(* Logix 5000 project; controller PLC_MCC1300_75F1 vendor 1 type 14 code 166 rev 32.11; software revision 32.04; part 28 of 83 *)
(* tags used below, declared in another part *)
   AUX_tCapsConveyor_NULL : UDT_CapsConveyor_ZC;
   AUX_xInitialize : BOOL;
   CM_AreaStackerToLine_JS1 : CM_AreaStackerToLine;
   CM_AreaStackerToLine_JS1_Sync : CM_AreaStackerToLine;
   CM_AreaStackerToLine_JS2 : CM_AreaStackerToLine;
   CM_AreaStackerToLine_JS2_Sync : CM_AreaStackerToLine;
   CM_ConveyorStackerToLine_JS1 : CM_ConveyorStackerToLine;
   CM_ConveyorStackerToLine_JS1_Sync : CM_ConveyorStackerToLine;
   CM_ConveyorStackerToLine_JS2 : CM_ConveyorStackerToLine;
   CM_ConveyorStackerToLine_JS2_Sync : CM_ConveyorStackerToLine;
   CM_DATA_Z410_Rx : UDT_PlateData_Convoy;
   CM_DATA_Z410_Rx_Sync : UDT_PlateData_Convoy;
   CM_DATA_Z410_Rx_TmpBuffer : SINT[104];
   CM_DATA_Z410_Tx : UDT_PlateData_Convoy;
   CM_DATA_Z410_Tx_MSG : MESSAGE;
   CM_DATA_Z410_Tx_PH : DINT;
   CM_DATA_Z410_Tx_TempBuffer : SINT[104];
   CM_DATA_Z410_Tx_tmON : TIMER;
   CM_DATA_Z420_Rx : UDT_PlateData_Convoy;
   CM_DATA_Z420_Rx_Sync : UDT_PlateData_Convoy;
   CM_DATA_Z420_Rx_TmpBuffer : SINT[104];
   CM_DATA_Z420_Tx : UDT_PlateData_Convoy;
   CM_DATA_Z420_Tx_MSG : MESSAGE;
   CM_DATA_Z420_Tx_PH : DINT;
   CM_DATA_Z420_Tx_TempBuffer : SINT[104];
   CM_DATA_Z420_Tx_tmON : TIMER;
   CM_LineToAreaStacker_JS1 : CM_LineToAreaStacker;
   CM_LineToAreaStacker_JS2 : CM_LineToAreaStacker;
   CM_LineToConveyorStacker_JS1 : CM_LineToConveyorStacker;
   CM_LineToConveyorStacker_JS2 : CM_LineToConveyorStacker;
   CNV10_FLT : ALIAS FOR I[4].9;
   CNV11_FLT : ALIAS FOR I[4].10;
   CNV12_FLT : ALIAS FOR I[4].11;
   CNV1_FLT : ALIAS FOR I[4].0;
   CNV2_FLT : ALIAS FOR I[4].1;
   CNV3_FLT : ALIAS FOR I[4].2;
   CNV4_FLT : ALIAS FOR I[4].3;
   CNV5_FLT : ALIAS FOR I[4].4;
   CNV6_FLT : ALIAS FOR I[4].5;
   CNV7_FLT : ALIAS FOR I[4].6;
   CNV8_FLT : ALIAS FOR I[4].7;
   CNV9_FLT : ALIAS FOR I[4].8;
   CONST_tPlant : UDT_PLANT_CONSTANTS;
   DROP_NO1_CRSH : ALIAS FOR I[73].12;
   GP_OB_InitializeMain : GP_OB_Initialize;
   GP_OB_InitializeMain_STC : GP_OB_Initialize_STC;
   I : INT[128];   // Local Input Updates Input Slot 2
   M2_DRV_CONT_ON : ALIAS FOR I[2].1;
   M2_DRV_FLT_LMP : ALIAS FOR O[9].0;
   M302SpeedUp : MAC_SpeedUp;
   M307ASpeedUp : MAC_SpeedUp;
   M30xTrimDeck : MAC_TrimmingDeck[5];
   M30xTrimWheel : MAC_TrimmingWheels[5];
   M310Popup : MAC_Popup_ZC[2];
   M310Popup_SL_DATA : UDT_Convoy_SL;
   M312 : MAC_Conveyor_Single;
   M312_SpaceConv_Utilities : SpaceConv_Utilities;
   M315Popup : MAC_Popup_ZC[2];
   M315Popup_SL_DATA : UDT_Convoy_SL;
   M350Popup : MAC_Popup_ZC;
   M410_DATA_xSendERR : BOOL;
   M420_DATA_xSendERR : BOOL;
   N130 : INT[8];
   N131 : INT[8];
   O : INT[128];
   REL_DATARCVD_N : ALIAS FOR O[54].2;
   REL_DATARCVDS : ALIAS FOR O[58].2;
   REL_REJWINLAMPN : ALIAS FOR O[54].3;
   REL_REJWINLAMPS : ALIAS FOR O[58].3;
   T4 : TIMER[51];
   TMP_d : DINT;
   TMP_dIndex : DINT;
   TMP_dIndexCapConv : DINT;
   TMP_dIndexConv : DINT;
   TMP_dLineSize : DINT;
   tony_always_false : BOOL;
   xAlwaysOFF : BOOL;
   Z300_Conveyor : UDT_StandConv[29];
   Z300_Conveyor_Conf : UDT_Conveyor_Config[29];
   Z300_dEndTrackingPosition : DINT;
   Z300_dStartTrackingPosition : DINT;
   Z300_LineTracking : UDT_LINE_TRACKING;
   Z301 : MAC_Zone_ML;
   Z401 : MAC_Zone;
   Z401_HMW : MAC_Zone_HMW;

PROGRAM Communication   (* main routine Main *)

ROUTINE CM_Z410   (* ladder *)
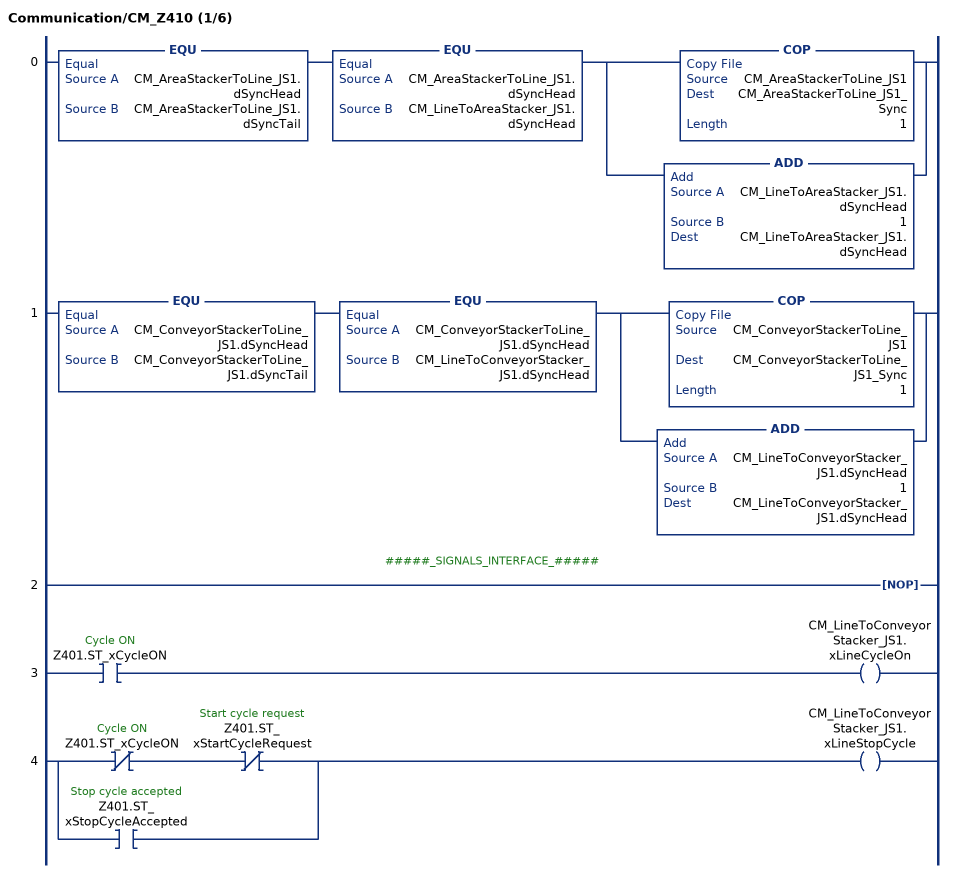
   0: EQU(CM_AreaStackerToLine_JS1.dSyncHead,CM_AreaStackerToLine_JS1.dSyncTail)EQU(CM_AreaStackerToLine_JS1.dSyncHead,CM_LineToAreaStacker_JS1.dSyncHead)[COP(CM_AreaStackerToLine_JS1,CM_AreaStackerToLine_JS1_Sync,1) ,ADD(CM_LineToAreaStacker_JS1.dSyncHead,1,CM_LineToAreaStacker_JS1.dSyncHead) ];
   1: EQU(CM_ConveyorStackerToLine_JS1.dSyncHead,CM_ConveyorStackerToLine_JS1.dSyncTail)EQU(CM_ConveyorStackerToLine_JS1.dSyncHead,CM_LineToConveyorStacker_JS1.dSyncHead)[COP(CM_ConveyorStackerToLine_JS1,CM_ConveyorStackerToLine_JS1_Sync,1) ,ADD(CM_LineToConveyorStacker_JS1.dSyncHead,1,CM_LineToConveyorStacker_JS1.dSyncHead) ];
   // #####_SIGNALS_INTERFACE_#####
   2: NOP();
   3: XIC(Z401.ST_xCycleON)OTE(CM_LineToConveyorStacker_JS1.xLineCycleOn);
   4: [XIO(Z401.ST_xCycleON) XIO(Z401.ST_xStartCycleRequest) ,XIC(Z401.ST_xStopCycleAccepted) ]OTE(CM_LineToConveyorStacker_JS1.xLineStopCycle);
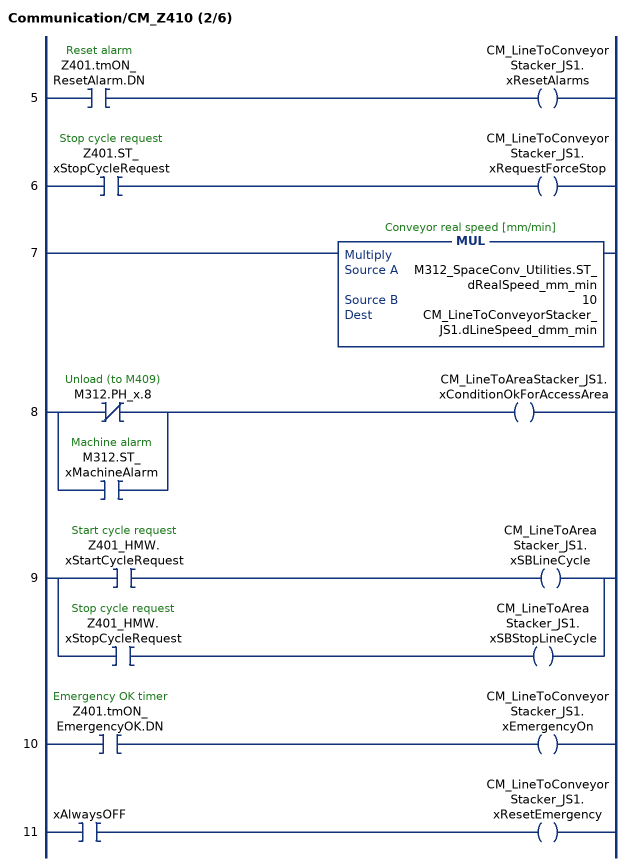
   5: XIC(Z401.tmON_ResetAlarm.DN)OTE(CM_LineToConveyorStacker_JS1.xResetAlarms);
   6: XIC(Z401.ST_xStopCycleRequest)OTE(CM_LineToConveyorStacker_JS1.xRequestForceStop);
   7: MUL(M312_SpaceConv_Utilities.ST_dRealSpeed_mm_min,10,CM_LineToConveyorStacker_JS1.dLineSpeed_dmm_min);
   8: [XIO(M312.PH_x.8) ,XIC(M312.ST_xMachineAlarm) ]OTE(CM_LineToAreaStacker_JS1.xConditionOkForAccessArea);
   9: [XIC(Z401_HMW.xStartCycleRequest) OTE(CM_LineToAreaStacker_JS1.xSBLineCycle) ,XIC(Z401_HMW.xStopCycleRequest) OTE(CM_LineToAreaStacker_JS1.xSBStopLineCycle) ];
   10: XIC(Z401.tmON_EmergencyOK.DN)OTE(CM_LineToConveyorStacker_JS1.xEmergencyOn);
   11: XIC(xAlwaysOFF)OTE(CM_LineToConveyorStacker_JS1.xResetEmergency);
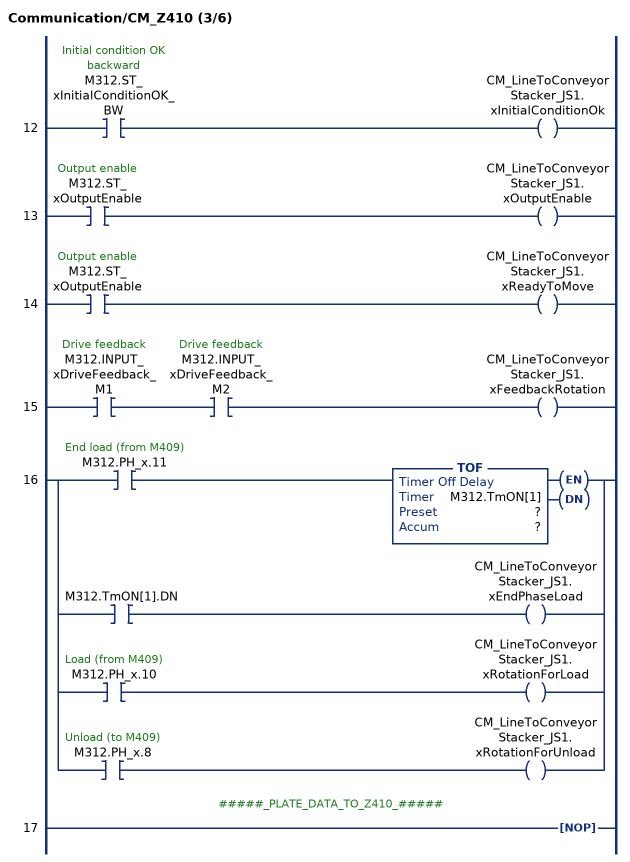
   12: XIC(M312.ST_xInitialConditionOK_BW)OTE(CM_LineToConveyorStacker_JS1.xInitialConditionOk);
   13: XIC(M312.ST_xOutputEnable)OTE(CM_LineToConveyorStacker_JS1.xOutputEnable);
   14: XIC(M312.ST_xOutputEnable)OTE(CM_LineToConveyorStacker_JS1.xReadyToMove);
   15: XIC(M312.INPUT_xDriveFeedback_M1)XIC(M312.INPUT_xDriveFeedback_M2)OTE(CM_LineToConveyorStacker_JS1.xFeedbackRotation);
   16: [[XIC(M312.PH_x.11) TOF(M312.TmON[1],?,?) ,XIC(M312.TmON[1].DN) OTE(CM_LineToConveyorStacker_JS1.xEndPhaseLoad) ] ,XIC(M312.PH_x.10) OTE(CM_LineToConveyorStacker_JS1.xRotationForLoad) ,XIC(M312.PH_x.8) OTE(CM_LineToConveyorStacker_JS1.xRotationForUnload) ];
   // #####_PLATE_DATA_TO_Z410_#####
   17: NOP();
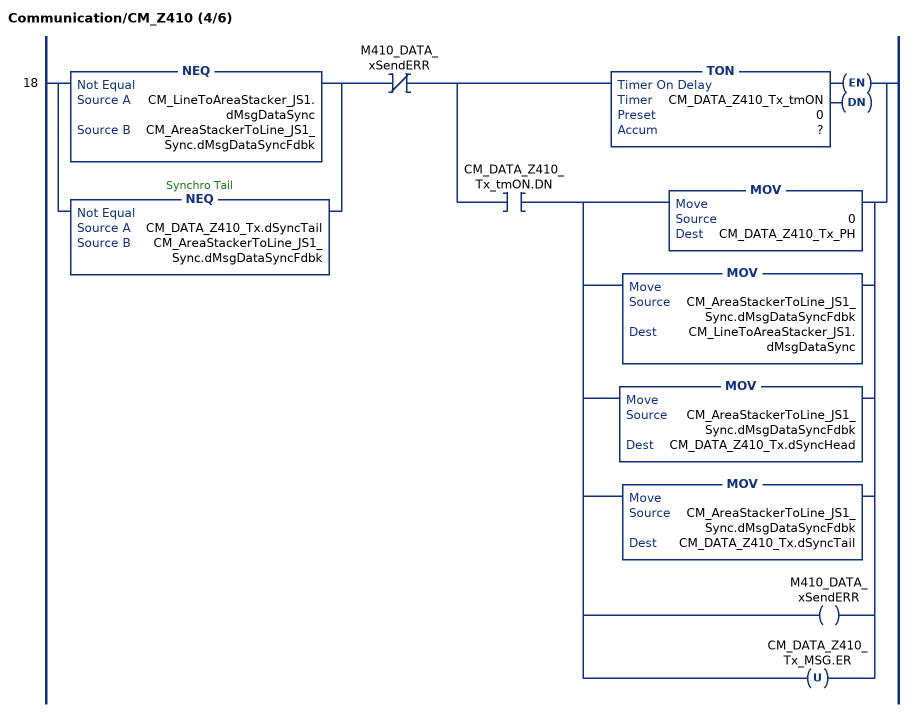
   18: [NEQ(CM_LineToAreaStacker_JS1.dMsgDataSync,CM_AreaStackerToLine_JS1_Sync.dMsgDataSyncFdbk) ,NEQ(CM_DATA_Z410_Tx.dSyncTail,CM_AreaStackerToLine_JS1_Sync.dMsgDataSyncFdbk) ]XIO(M410_DATA_xSendERR)[TON(CM_DATA_Z410_Tx_tmON,?,?) ,XIC(CM_DATA_Z410_Tx_tmON.DN) [MOV(0,CM_DATA_Z410_Tx_PH) ,MOV(CM_AreaStackerToLine_JS1_Sync.dMsgDataSyncFdbk,CM_LineToAreaStacker_JS1.dMsgDataSync) ,MOV(CM_AreaStackerToLine_JS1_Sync.dMsgDataSyncFdbk,CM_DATA_Z410_Tx.dSyncHead) ,MOV(CM_AreaStackerToLine_JS1_Sync.dMsgDataSyncFdbk,CM_DATA_Z410_Tx.dSyncTail) ,OTE(M410_DATA_xSendERR) ,OTU(CM_DATA_Z410_Tx_MSG.ER) ] ];
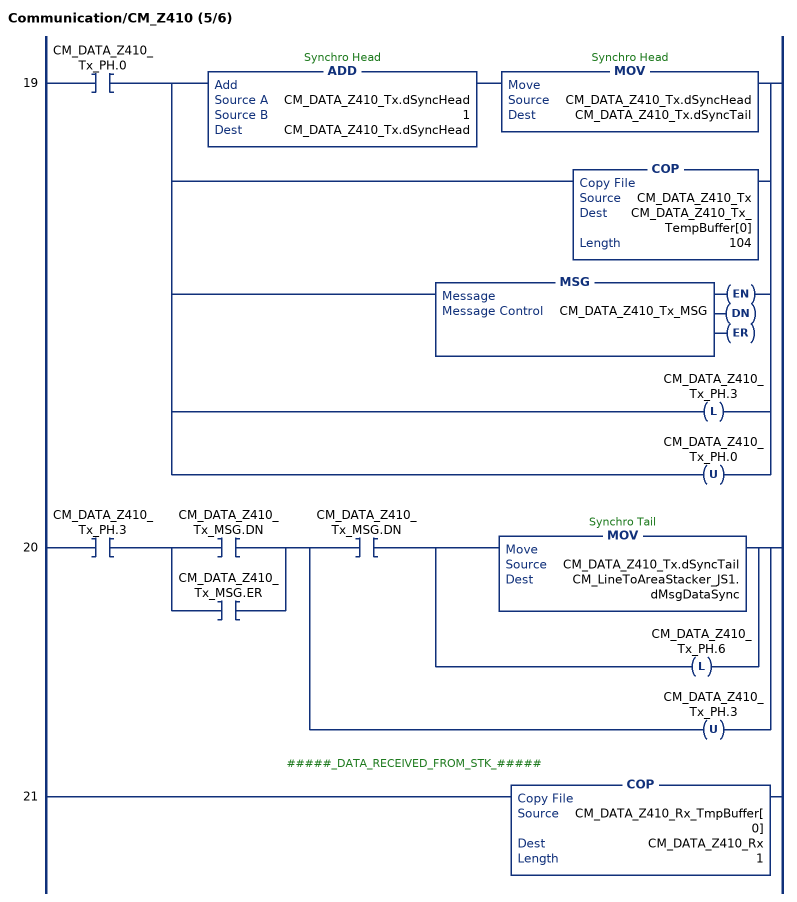
   19: XIC(CM_DATA_Z410_Tx_PH.0)[ADD(CM_DATA_Z410_Tx.dSyncHead,1,CM_DATA_Z410_Tx.dSyncHead) MOV(CM_DATA_Z410_Tx.dSyncHead,CM_DATA_Z410_Tx.dSyncTail) ,COP(CM_DATA_Z410_Tx,CM_DATA_Z410_Tx_TempBuffer[0],104) ,MSG(CM_DATA_Z410_Tx_MSG) ,OTL(CM_DATA_Z410_Tx_PH.3) ,OTU(CM_DATA_Z410_Tx_PH.0) ];
   20: XIC(CM_DATA_Z410_Tx_PH.3)[XIC(CM_DATA_Z410_Tx_MSG.DN) ,XIC(CM_DATA_Z410_Tx_MSG.ER) ][XIC(CM_DATA_Z410_Tx_MSG.DN) [MOV(CM_DATA_Z410_Tx.dSyncTail,CM_LineToAreaStacker_JS1.dMsgDataSync) ,OTL(CM_DATA_Z410_Tx_PH.6) ] ,OTU(CM_DATA_Z410_Tx_PH.3) ];
   // #####_DATA_RECEIVED_FROM_STK_#####
   21: COP(CM_DATA_Z410_Rx_TmpBuffer[0],CM_DATA_Z410_Rx,1);
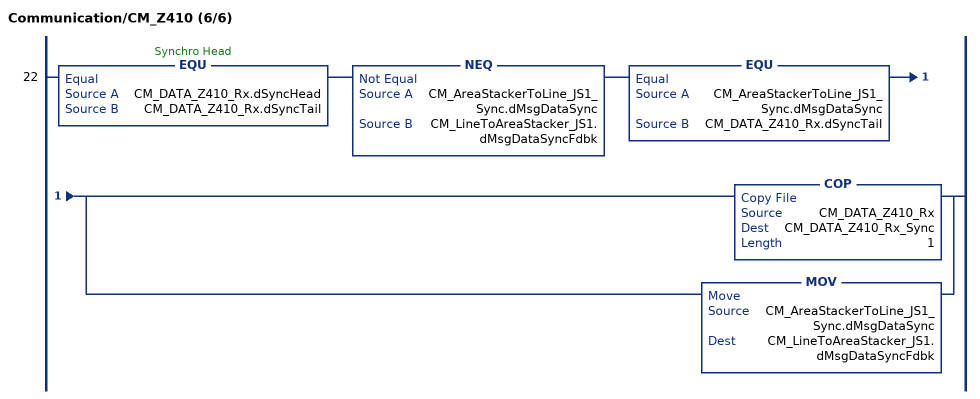
   22: EQU(CM_DATA_Z410_Rx.dSyncHead,CM_DATA_Z410_Rx.dSyncTail)NEQ(CM_AreaStackerToLine_JS1_Sync.dMsgDataSync,CM_LineToAreaStacker_JS1.dMsgDataSyncFdbk)EQU(CM_AreaStackerToLine_JS1_Sync.dMsgDataSync,CM_DATA_Z410_Rx.dSyncTail)[COP(CM_DATA_Z410_Rx,CM_DATA_Z410_Rx_Sync,1) ,MOV(CM_AreaStackerToLine_JS1_Sync.dMsgDataSync,CM_LineToAreaStacker_JS1.dMsgDataSyncFdbk) ];
END_ROUTINE

ROUTINE CM_Z420   (* ladder *)
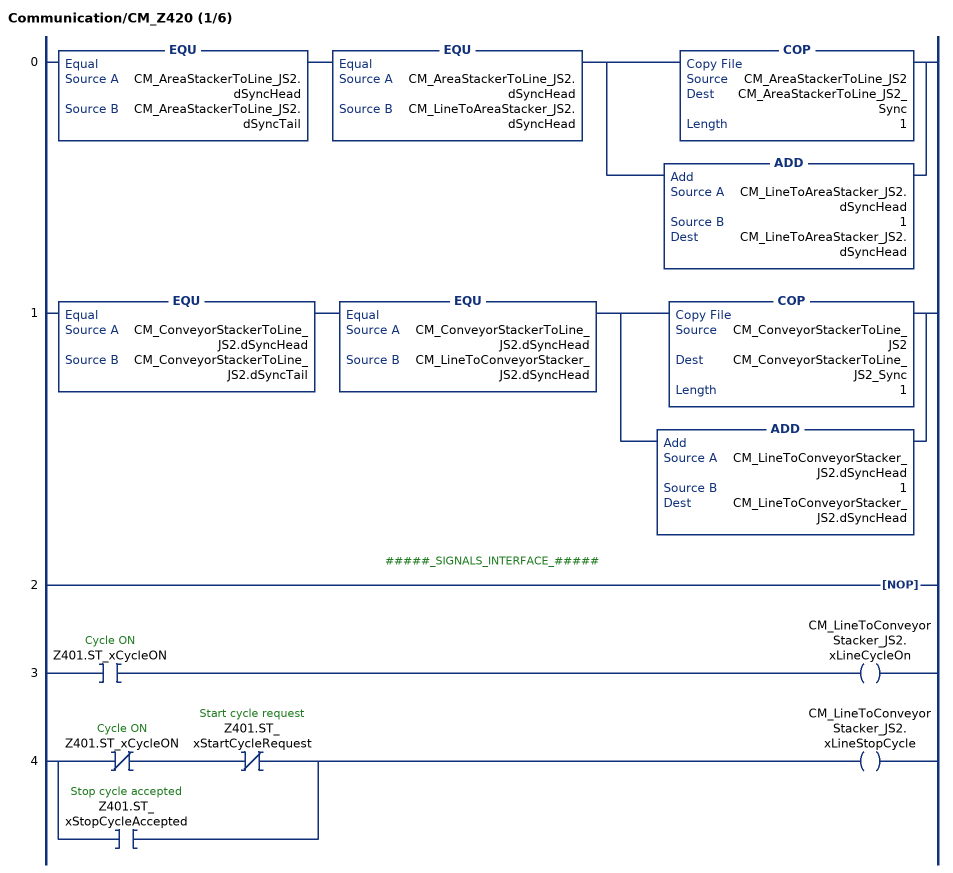
   0: EQU(CM_AreaStackerToLine_JS2.dSyncHead,CM_AreaStackerToLine_JS2.dSyncTail)EQU(CM_AreaStackerToLine_JS2.dSyncHead,CM_LineToAreaStacker_JS2.dSyncHead)[COP(CM_AreaStackerToLine_JS2,CM_AreaStackerToLine_JS2_Sync,1) ,ADD(CM_LineToAreaStacker_JS2.dSyncHead,1,CM_LineToAreaStacker_JS2.dSyncHead) ];
   1: EQU(CM_ConveyorStackerToLine_JS2.dSyncHead,CM_ConveyorStackerToLine_JS2.dSyncTail)EQU(CM_ConveyorStackerToLine_JS2.dSyncHead,CM_LineToConveyorStacker_JS2.dSyncHead)[COP(CM_ConveyorStackerToLine_JS2,CM_ConveyorStackerToLine_JS2_Sync,1) ,ADD(CM_LineToConveyorStacker_JS2.dSyncHead,1,CM_LineToConveyorStacker_JS2.dSyncHead) ];
   // #####_SIGNALS_INTERFACE_#####
   2: NOP();
   3: XIC(Z401.ST_xCycleON)OTE(CM_LineToConveyorStacker_JS2.xLineCycleOn);
   4: [XIO(Z401.ST_xCycleON) XIO(Z401.ST_xStartCycleRequest) ,XIC(Z401.ST_xStopCycleAccepted) ]OTE(CM_LineToConveyorStacker_JS2.xLineStopCycle);
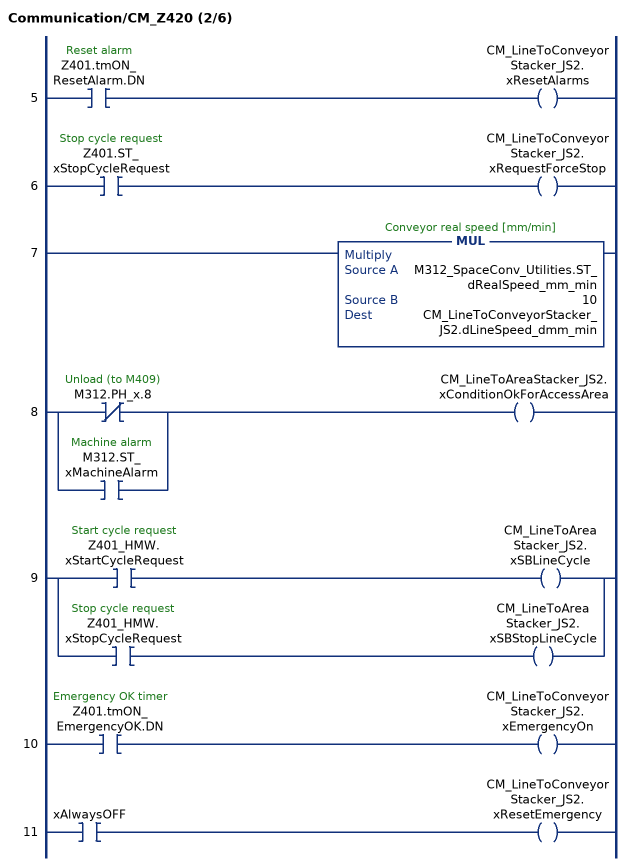
   5: XIC(Z401.tmON_ResetAlarm.DN)OTE(CM_LineToConveyorStacker_JS2.xResetAlarms);
   6: XIC(Z401.ST_xStopCycleRequest)OTE(CM_LineToConveyorStacker_JS2.xRequestForceStop);
   7: MUL(M312_SpaceConv_Utilities.ST_dRealSpeed_mm_min,10,CM_LineToConveyorStacker_JS2.dLineSpeed_dmm_min);
   8: [XIO(M312.PH_x.8) ,XIC(M312.ST_xMachineAlarm) ]OTE(CM_LineToAreaStacker_JS2.xConditionOkForAccessArea);
   9: [XIC(Z401_HMW.xStartCycleRequest) OTE(CM_LineToAreaStacker_JS2.xSBLineCycle) ,XIC(Z401_HMW.xStopCycleRequest) OTE(CM_LineToAreaStacker_JS2.xSBStopLineCycle) ];
   10: XIC(Z401.tmON_EmergencyOK.DN)OTE(CM_LineToConveyorStacker_JS2.xEmergencyOn);
   11: XIC(xAlwaysOFF)OTE(CM_LineToConveyorStacker_JS2.xResetEmergency);
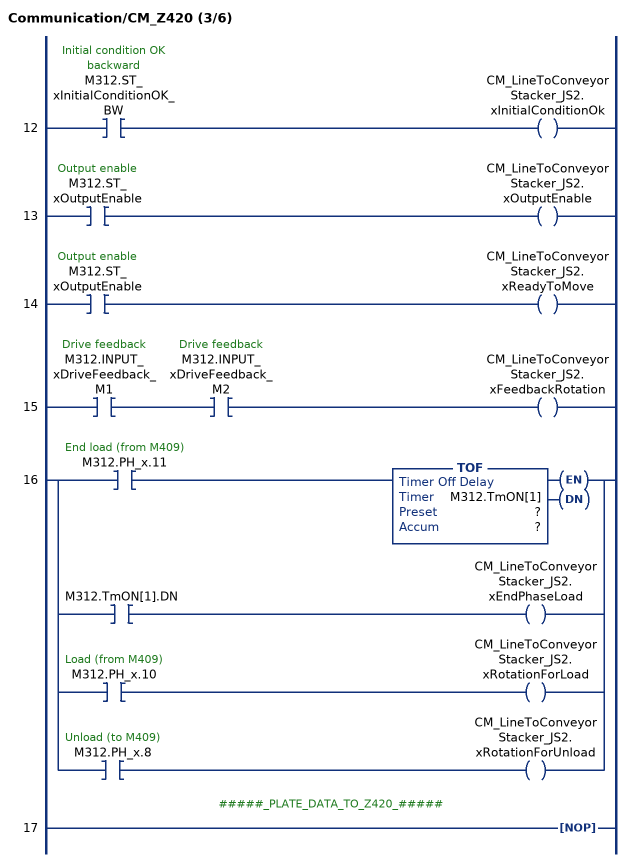
   12: XIC(M312.ST_xInitialConditionOK_BW)OTE(CM_LineToConveyorStacker_JS2.xInitialConditionOk);
   13: XIC(M312.ST_xOutputEnable)OTE(CM_LineToConveyorStacker_JS2.xOutputEnable);
   14: XIC(M312.ST_xOutputEnable)OTE(CM_LineToConveyorStacker_JS2.xReadyToMove);
   15: XIC(M312.INPUT_xDriveFeedback_M1)XIC(M312.INPUT_xDriveFeedback_M2)OTE(CM_LineToConveyorStacker_JS2.xFeedbackRotation);
   16: [[XIC(M312.PH_x.11) TOF(M312.TmON[1],?,?) ,XIC(M312.TmON[1].DN) OTE(CM_LineToConveyorStacker_JS2.xEndPhaseLoad) ] ,XIC(M312.PH_x.10) OTE(CM_LineToConveyorStacker_JS2.xRotationForLoad) ,XIC(M312.PH_x.8) OTE(CM_LineToConveyorStacker_JS2.xRotationForUnload) ];
   // #####_PLATE_DATA_TO_Z420_#####
   17: NOP();
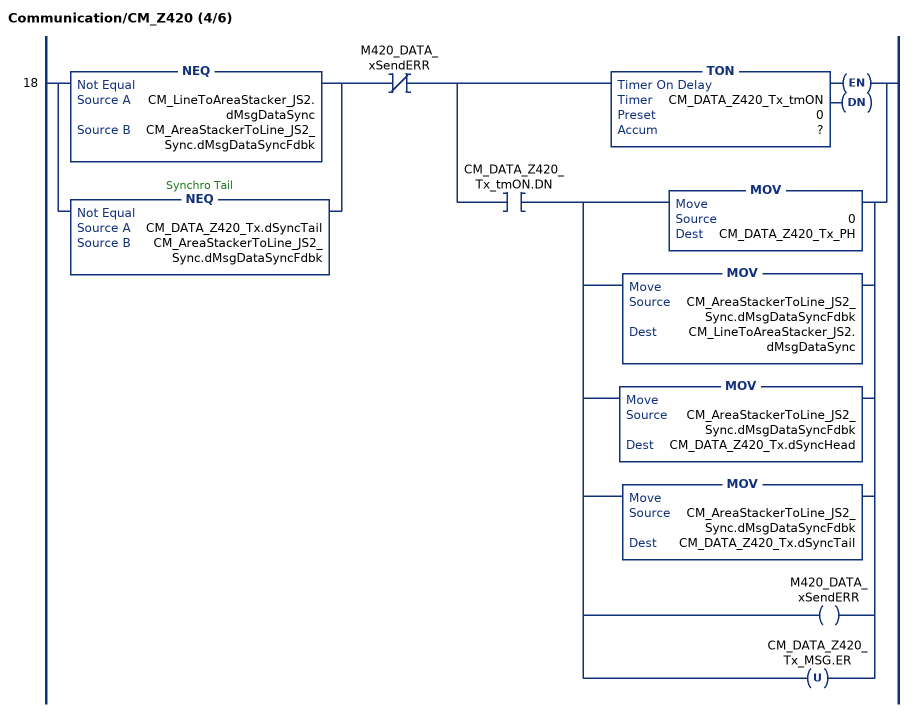
   18: [NEQ(CM_LineToAreaStacker_JS2.dMsgDataSync,CM_AreaStackerToLine_JS2_Sync.dMsgDataSyncFdbk) ,NEQ(CM_DATA_Z420_Tx.dSyncTail,CM_AreaStackerToLine_JS2_Sync.dMsgDataSyncFdbk) ]XIO(M420_DATA_xSendERR)[TON(CM_DATA_Z420_Tx_tmON,?,?) ,XIC(CM_DATA_Z420_Tx_tmON.DN) [MOV(0,CM_DATA_Z420_Tx_PH) ,MOV(CM_AreaStackerToLine_JS2_Sync.dMsgDataSyncFdbk,CM_LineToAreaStacker_JS2.dMsgDataSync) ,MOV(CM_AreaStackerToLine_JS2_Sync.dMsgDataSyncFdbk,CM_DATA_Z420_Tx.dSyncHead) ,MOV(CM_AreaStackerToLine_JS2_Sync.dMsgDataSyncFdbk,CM_DATA_Z420_Tx.dSyncTail) ,OTE(M420_DATA_xSendERR) ,OTU(CM_DATA_Z420_Tx_MSG.ER) ] ];
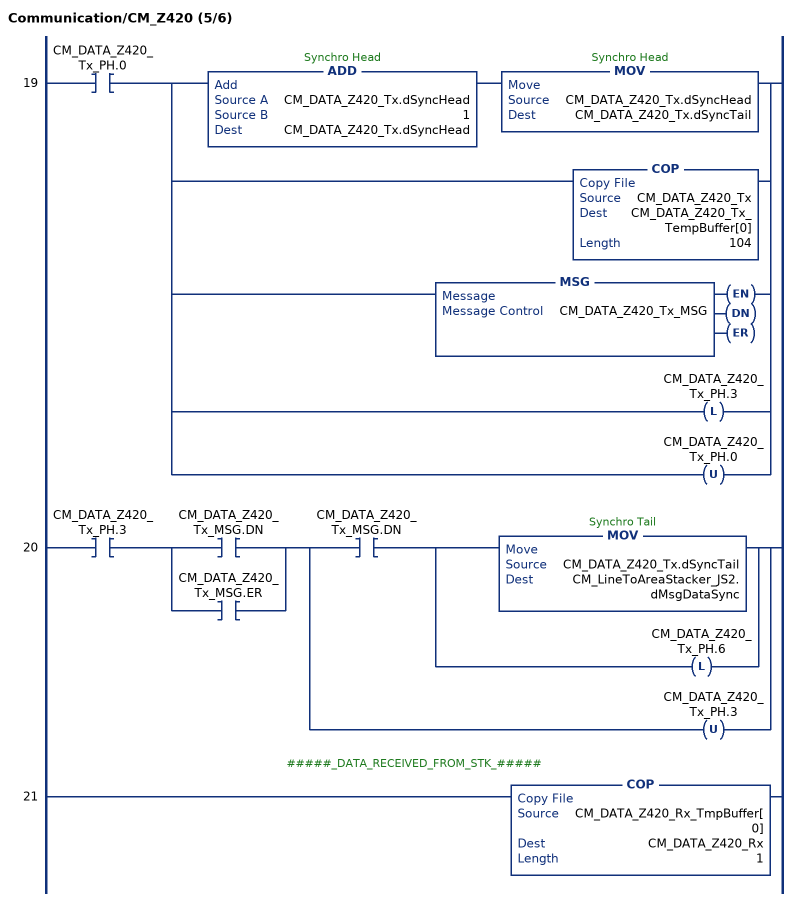
   19: XIC(CM_DATA_Z420_Tx_PH.0)[ADD(CM_DATA_Z420_Tx.dSyncHead,1,CM_DATA_Z420_Tx.dSyncHead) MOV(CM_DATA_Z420_Tx.dSyncHead,CM_DATA_Z420_Tx.dSyncTail) ,COP(CM_DATA_Z420_Tx,CM_DATA_Z420_Tx_TempBuffer[0],104) ,MSG(CM_DATA_Z420_Tx_MSG) ,OTL(CM_DATA_Z420_Tx_PH.3) ,OTU(CM_DATA_Z420_Tx_PH.0) ];
   20: XIC(CM_DATA_Z420_Tx_PH.3)[XIC(CM_DATA_Z420_Tx_MSG.DN) ,XIC(CM_DATA_Z420_Tx_MSG.ER) ][XIC(CM_DATA_Z420_Tx_MSG.DN) [MOV(CM_DATA_Z420_Tx.dSyncTail,CM_LineToAreaStacker_JS2.dMsgDataSync) ,OTL(CM_DATA_Z420_Tx_PH.6) ] ,OTU(CM_DATA_Z420_Tx_PH.3) ];
   // #####_DATA_RECEIVED_FROM_STK_#####
   21: COP(CM_DATA_Z420_Rx_TmpBuffer[0],CM_DATA_Z420_Rx,1);
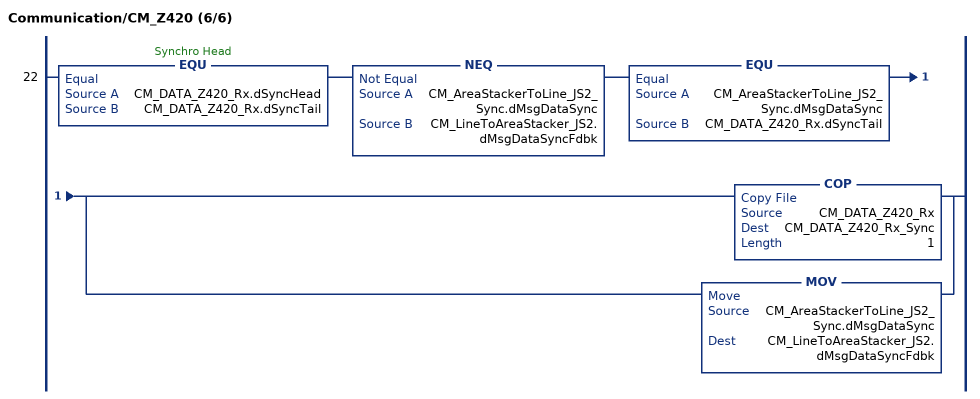
   22: EQU(CM_DATA_Z420_Rx.dSyncHead,CM_DATA_Z420_Rx.dSyncTail)NEQ(CM_AreaStackerToLine_JS2_Sync.dMsgDataSync,CM_LineToAreaStacker_JS2.dMsgDataSyncFdbk)EQU(CM_AreaStackerToLine_JS2_Sync.dMsgDataSync,CM_DATA_Z420_Rx.dSyncTail)[COP(CM_DATA_Z420_Rx,CM_DATA_Z420_Rx_Sync,1) ,MOV(CM_AreaStackerToLine_JS2_Sync.dMsgDataSync,CM_LineToAreaStacker_JS2.dMsgDataSyncFdbk) ];
END_ROUTINE

ROUTINE Main   (* ladder *)